// TIA Portal project "HEAT-1-CADIZ-V16" (V20)

(* hardware
DEVICE "S7-1200 station_1"  S7-1200 Station
   slot 0: "Rack_0"  S7-1200 Rack  Rack  V1.0
   slot 1: "PLC_1"  CPU 1214FC DC/DC/RLY  6ES7 214-1HF40-0XB0  V4.6
   slot 2: "DI 16x24VDC_1"  6ES7 221-1BH32-0XB0  V2.0
   slot 3: "DQ 16xRelay_1"  SM 1222 DQ16 x relay  6ES7 222-1HH32-0XB0  V2.0
   slot 4: "F-DI 8/16x24VDC_1"  SM 1226 F-DI8/16 x 24VDC  6ES7 226-6BA32-0XB0  V2.0
   slot 5: "F-DI 8/16x24VDC_2"  SM 1226 F-DI8/16 x 24VDC  6ES7 226-6BA32-0XB0  V2.0
   slot 6: "F-DQ 4x24VDC_1"  SM 1226 F-DQ4 x 24VDC  6ES7 226-6DA32-0XB0  V2.0
DEVICE "GSD device_1"  GSD.Device.PN
   slot 0: "Rack"  Rack  V1.0
   slot 0: "KRC5"  KUKA.PROFINET 6.0  0x300  V6.0
      slot 0: "KUKA.PROFINET 6.0"  KUKA.PROFINET 6.0
      slot 1: "Interface1"  Interface1
         slot 1: "Port001(XF3)"  Port001(XF3)
         slot 2: "Port002(XF4)"  Port002(XF4)
         slot 3: "Port003(XF5)"  Port003(XF5)
         slot 4: "Port004(XF6)"  Port004(XF6)
   slot 1: "64 safe digital in- and outputs (2.4)_1"  64 safe digital in- and outputs (2.4)  KUKADevF64_2.4
      slot 0: "64 safe digital in- and outputs (2.4)"  64 safe digital in- and outputs (2.4)
   slot 2: "512 digital in- and outputs_1"  512 digital in- and outputs  KUKA Device IO512
      slot 0: "512 digital in- and outputs"  512 digital in- and outputs
DEVICE "HMI_1"  KTP1200 Basic PN
   slot 0: "HMI_1"  KTP1200 Basic PN  6AV2 123-2MB03-0AX0  17.0.0.0
   slot 1: "HMI_RT_1"  KTP1200 Basic PN  6AV2 123-2MB03-0AX0  17.0.0.0
   slot 5: "HMI_1.IE_CP_1"  PROFINET Interface  17.0.0.0
      slot 1: "PROFINET Interface_1"  PROFINET Interface
         slot 1: "Port_1"  Port
DEVICE "ET 200SP station_2"  ET 200SP-Station
   slot 0: "Rack_0"  Rack  6ES5 710-8MAx1
   slot 0: "islaparking"  IM 155-6 PN ST  6ES7 155-6AU01-0BN0  V4.2
   slot 1: "DI 16x24VDC ST_1"  DI 16x24VDC ST  6ES7 131-6BH01-0BA0  V0.0
      slot 1: "DI 16x24VDC ST_1"  DI 16x24VDC ST
   slot 2: "DI 8x24VDC ST_1"  DI 8x24VDC ST  6ES7 131-6BF01-0BA0  V0.0
      slot 1: "DI 8x24VDC ST_1"  DI 8x24VDC ST
   slot 3: "DQ 16x24VDC/0.5A ST_1"  DQ 16x24VDC/0.5A ST  6ES7 132-6BH01-0BA0  V0.0
      slot 1: "DQ 16x24VDC/0.5A ST_1"  DQ 16x24VDC/0.5A ST
   slot 4: "DQ 8x24VDC/0.5A ST_1"  DQ 8x24VDC/0.5A ST  6ES7 132-6BF01-0BA0  V0.0
      slot 1: "DQ 8x24VDC/0.5A ST_1"  DQ 8x24VDC/0.5A ST
   slot 5: "Server module_1"  Server module  6ES7 193-6PA00-0AA0  V1.1
      slot 1: "Server module_1"  Server module
   slot 127: "BA 2xRJ45"  BA 2xRJ45  6ES7 193-6AR00-0AA0  V0.0
      slot 1: "Port_1"  X1 P1R  6ES7 193-6AR00-0AA0  V0.0
      slot 2: "Port_2"  X1 P2R  6ES7 193-6AR00-0AA0  V0.0
DEVICE "ET 200SP station_1"  ET 200SP-Station
   slot 0: "Rack_0"  Rack  6ES5 710-8MAx1
   slot 0: "islarobot"  IM 155-6 PN ST  6ES7 155-6AU01-0BN0  V4.2
   slot 1: "DI 16x24VDC ST_1"  DI 16x24VDC ST  6ES7 131-6BH01-0BA0  V0.0
      slot 1: "DI 16x24VDC ST_1"  DI 16x24VDC ST
   slot 2: "DI 8x24VDC ST_1"  DI 8x24VDC ST  6ES7 131-6BF01-0BA0  V0.0
      slot 1: "DI 8x24VDC ST_1"  DI 8x24VDC ST
   slot 3: "DQ 16x24VDC/0.5A ST_1"  DQ 16x24VDC/0.5A ST  6ES7 132-6BH01-0BA0  V0.0
      slot 1: "DQ 16x24VDC/0.5A ST_1"  DQ 16x24VDC/0.5A ST
   slot 4: "DQ 8x24VDC/0.5A ST_1"  DQ 8x24VDC/0.5A ST  6ES7 132-6BF01-0BA0  V0.0
      slot 1: "DQ 8x24VDC/0.5A ST_1"  DQ 8x24VDC/0.5A ST
   slot 5: "Server module_1"  Server module  6ES7 193-6PA00-0AA0  V1.1
      slot 1: "Server module_1"  Server module
   slot 127: "BA 2xRJ45"  BA 2xRJ45  6ES7 193-6AR00-0AA0  V0.0
      slot 1: "Port_1"  X1 P1R  6ES7 193-6AR00-0AA0  V0.0
      slot 2: "Port_2"  X1 P2R  6ES7 193-6AR00-0AA0  V0.0
DEVICE "GSD device_2"  GSD.Device.PN
   slot 0: "Rack"  Rack  V1.0
   slot 0: "CPX"  CPX Rev 50  TN 197330
      slot 0: "CPX Rev 50"  CPX Rev 50
      slot 1: "PN-IO Interface"  PN-IO Interface
         slot 1: "Port 1"  Port 1
         slot 2: "Port 2"  Port 2
   slot 1: "FB43 PNIO Module_1"  FB43 PNIO Module  TN 8110369, CPX-FB43
      slot 0: "FB43 PNIO Module"  FB43 PNIO Module
   slot 2: "MPAL DIL 4 [32DO]_1"  MPAL DIL 4 [32DO]
      slot 0: "MPAL DIL 4 [32DO]"  MPAL DIL 4 [32DO]
DEVICE "ET 200SP station_3"  ET 200SP-Station
   slot 0: "Rack_0"  Rack  6ES5 710-8MAx1
   slot 0: "sistemadeagua"  IM 155-6 PN ST  6ES7 155-6AU01-0BN0  V4.2
   slot 1: "DI 8x24VDC ST_1"  DI 8x24VDC ST  6ES7 131-6BF01-0BA0  V0.0
      slot 1: "DI 8x24VDC ST_1"  DI 8x24VDC ST
   slot 2: "DQ 8x24VDC/0.5A ST_1"  DQ 8x24VDC/0.5A ST  6ES7 132-6BF01-0BA0  V0.0
      slot 1: "DQ 8x24VDC/0.5A ST_1"  DQ 8x24VDC/0.5A ST
   slot 3: "AI 4xU/I 2-wire ST_1"  AI 4xU/I 2-wire ST  6ES7 134-6HD01-0BA1  V2.0
      slot 1: "AI 4xU/I 2-wire ST_1"  AI 4xU/I 2-wire ST
   slot 4: "Server module_1"  Server module  6ES7 193-6PA00-0AA0  V1.1
      slot 1: "Server module_1"  Server module
   slot 127: "BA 2xRJ45"  BA 2xRJ45  6ES7 193-6AR00-0AA0  V0.0
      slot 1: "Port_1"  X1 P1R  6ES7 193-6AR00-0AA0  V0.0
      slot 2: "Port_2"  X1 P2R  6ES7 193-6AR00-0AA0  V0.0
*)

// ===== PLC "PLC_1"  CPU 1214FC DC/DC/RLY =====

VAR_GLOBAL   // PLC tag table "Default tag table"
   "RES1 (reservado)" AT %Q500.0 : Bool;
   "eStopButtonCabinet" AT %I40.0 : Bool;   // Emergency-Stop cabinet — 1oo2 result
   "eStopButtonTank" AT %I40.1 : Bool;   // Emergency-Stop tank — 1oo2 result
   "eStopButtonTankPartnerCh" AT %I41.1 : Bool;   // partner channel 1oo2 — do not use
   "eStopButtonWaterSystem" AT %I40.2 : Bool;   // Emergency-Stop water system — 1oo2 result
   "eStopButtonWaterSystemPartnerCh" AT %I41.2 : Bool;   // partner channel 1oo2 — do not use
   "eStopButtonHmiPanel" AT %I40.3 : Bool;   // Emergency-Stop HMI panel — 1oo2 result
   "eStopButtonHmiPanelPartnerCh" AT %I41.3 : Bool;   // partner channel 1oo2 — do not use
   "eStopButtonLightCurtain1" AT %I40.4 : Bool;   // Emergency-Stop light curtain 1 — 1oo2 resul
   "eStopButtonLightCurtain1PartnerCh" AT %I41.4 : Bool;   // partner channel 1oo2 — do not use
   "eStopButtonDoor" AT %I40.5 : Bool;   // Emergency-Stop Door — 1oo2 result
   "eStopButtonDoorPartnerCh" AT %I41.5 : Bool;   // partner channel 1oo2 — do not use
   "lightCurtain1Ossd1" AT %I50.0 : Bool;   // Z2 – LC 1 OSSD 1 (receiver)
   "lightCurtain1Ossd2" AT %I51.0 : Bool;   // Z2 – LC 1 OSSD 2 (receiver)
   "lightCurtain3Ossd1" AT %I50.1 : Bool;   // Z2 – LC 3 OSSD 1 (receiver)
   "lightCurtain3Ossd2" AT %I51.1 : Bool;   // Z2 – LC 3 OSSD 2 (receiver)
   "lightCurtain6Ossd1" AT %I50.2 : Bool;   // Z2 – LC 6 OSSD 1 (receiver)
   "lightCurtain6Ossd2" AT %I51.2 : Bool;   // Z2 – LC 6 OSSD 2 (receiver)
   "enableAccessReqSelector" AT %I50.3 : Bool;   // Rotary selector – enabless request access
   "DoorClosedCh1" AT %I50.6 : Bool;   // Safety door closed interlock – contact 1
   "resetDoorButton" AT %I50.7 : Bool;   // Reset push‑button
   "SAF_DOOR_CLSD_CH2" AT %I51.6 : Bool;   // Safety door closed interlock – contact 2
   "SAF_DOOR_UNLOCK_CH1" AT %Q60.0 : Bool;   // Unlock safety door – redundant output 1
   "SAF_GATE_UNLOCK_CH2" AT %Q60.2 : Bool;   // Unlock safety door – redundant output 2
   "IND_RESET_LAMP" AT %Q10.0 : Bool;   // Reset indicator lamp
   "IND_STATUS_LAMP" AT %Q10.1 : Bool;   // System-status pilot light
   "CMD_PRESS_EXH_VALVE" AT %Q11.0 : Bool;   // Pressure/exhaust solenoid-valve command
   "STS_RECIRC_PUMP" AT %I20.0 : Bool;   // Recirculation-pump feedback
   "STS_TRANSFER_PUMP" AT %I20.1 : Bool;   // Transfer-pump feedback
   "ALM_UV_FILTER" AT %I20.2 : Bool;   // UV-filter fault alarm
   "ALM_PIT_LVL_LOW" AT %I20.3 : Bool;   // Sump low-level alarm
   "ALM_TANK_LVL_LOW" AT %I20.4 : Bool;   // Tank low-level alarm
   "STS_TANK_FILLING" AT %I20.5 : Bool;   // Tank filling status
   "STS_TANK_DRAINING" AT %I20.6 : Bool;   // Tank draining status
   "MODE_WATER_AUTO" AT %Q30.3 : Bool;   // CONMUTADOR AUTO
   "IND_BEACON2_GREEN" AT %Q30.4 : Bool;   // Beacon 2 – green
   "IND_BEACON2_RED" AT %Q30.5 : Bool;   // Beacon 2 – red
   "robotPresenceSignalZone1" AT %I500.0 : Bool;
   "robotPresenceSignalZone2" AT %I500.1 : Bool;
   "robotPresenceSignalZone3" AT %I500.2 : Bool;
   "eStopButtonCabinetPartnerCh" AT %I41.0 : Bool;   // partner channel 1oo2 — do not use
   "lightCurtain2Ossd1" AT %I300.0 : Bool;
   "lightCurtain2Ossd2" AT %I301.0 : Bool;
   "eStopButtonIslandRightPartner" AT %I301.1 : Bool;
   "lightCurtain4Ossd1" AT %I350.0 : Bool;
   "eStopButtonIslandLeft" AT %I350.1 : Bool;
   "lightCurtain5Ossd1" AT %I350.2 : Bool;
   "eStopButtonIslandLefttPartner" AT %I350.3 : Bool;   // partner channel 1oo2 — do not use
   "lightCurtain4Ossd2" AT %I350.4 : Bool;
   "lightCurtain5Ossd2" AT %I350.6 : Bool;
   "accessReqButtonZone2" AT %I51.4 : Bool;   // Illuminated push-button – access request for zone 2
   "accessReqButtonZone3" AT %I51.5 : Bool;   // Illuminated push-button – access request for zone 3
   "accessReqButtonZone1" AT %I51.3 : Bool;   // Illuminated push-button – access request for zone 1
   "eStopButtonIslandRight" AT %I300.1 : Bool;
   "NHE – E‑Stop externo  NO pulsado" AT %Q500.1 : Bool;
   "BS – Puerta cerrada" AT %Q500.2 : Bool;
   "QBS – Ack puerta" AT %Q500.3 : Bool;
   "SHS1 – Stop 1" AT %Q500.4 : Bool;
   "SHS2 – Stop 2" AT %Q500.5 : Bool;
   "RES6" AT %Q500.6 : Bool;
   "RES7" AT %Q500.7 : Bool;
   "US2 – 24 V US2" AT %Q501.0 : Bool;
   "SBH – Safe Op Stop" AT %Q501.1 : Bool;
   "RES11" AT %Q501.2 : Bool;
   "RES12" AT %Q501.3 : Bool;
   "RES13" AT %Q501.4 : Bool;
   "RES14" AT %Q501.5 : Bool;
   "RES15" AT %Q501.6 : Bool;
   "SPA – Power‑down Ack" AT %Q501.7 : Bool;
   "resetHmiButton" AT %I51.7 : Bool;
   "Tag_1" AT %M200.0 : Bool;
   "Tag_2" AT %M201.0 : Bool;
   "Tag_3" AT %M500.1 : Bool;
   "Tag_4" AT %M755.5 : Bool;
   "V5" AT %Q0.4 : Bool;   // Biestable_B_RETROCESO
   "ABRIR_TAPA_PEPA" AT %Q170.2 : Bool;
   "CERRAR_TAPA_PEPA" AT %Q170.3 : Bool;
   "ABRIR_TAPA_INMERSION" AT %Q170.4 : Bool;
   "CERRAR_TAPA_INMERSION" AT %Q170.5 : Bool;
   "ABRIR_TAPA_MARCADOR" AT %Q170.6 : Bool;
   "CERRAR_TAPA_MARCADOR" AT %Q170.7 : Bool;
   "ABRIR_TAPA_PERFILOMETRO" AT %Q171.0 : Bool;
   "CERRAR_TAPA_PERFILOMETRO" AT %Q171.1 : Bool;
   "V6" AT %Q0.5 : Bool;   // Biestable_A_AVANCE
   "V7" AT %Q0.6 : Bool;
   "V8" AT %Q0.7 : Bool;
   "moveCode_00" AT %Q616.0 : Bool;
   "goTrigger" AT %Q622.0 : Bool;
   "baseReqId_00" AT %Q620.0 : Bool;
   "baseReqId_01" AT %Q620.1 : Bool;
   "baseReqId_02" AT %Q620.2 : Bool;
   "baseReqId_03" AT %Q620.3 : Bool;
   "baseReqId_04" AT %Q620.4 : Bool;
   "baseReqId_05" AT %Q620.5 : Bool;
   "baseReqId_06" AT %Q620.6 : Bool;
   "baseReqId_07" AT %Q620.7 : Bool;
   "baseReqId_08" AT %Q621.0 : Bool;
   "baseReqId_09" AT %Q621.1 : Bool;
   "baseReqId_10" AT %Q621.2 : Bool;
   "baseReqId_11" AT %Q621.3 : Bool;
   "baseReqId_12" AT %Q621.4 : Bool;
   "baseReqId_13" AT %Q621.5 : Bool;
   "baseReqId_14" AT %Q621.6 : Bool;
   "baseReqId_15" AT %Q621.7 : Bool;
   "moveCode_01" AT %Q616.1 : Bool;
   "moveCode_02" AT %Q616.2 : Bool;
   "moveCode_03" AT %Q616.3 : Bool;
   "moveCode_04" AT %Q616.4 : Bool;
   "moveCode_05" AT %Q616.5 : Bool;
   "moveCode_06" AT %Q616.6 : Bool;
   "moveCode_07" AT %Q616.7 : Bool;
   "moveCode_08" AT %Q617.0 : Bool;
   "moveCode_09" AT %Q617.1 : Bool;
   "moveCode_10" AT %Q617.2 : Bool;
   "moveCode_11" AT %Q617.3 : Bool;
   "moveCode_12" AT %Q617.4 : Bool;
   "moveCode_13" AT %Q617.5 : Bool;
   "moveCode_14" AT %Q617.6 : Bool;
   "moveCode_15" AT %Q617.7 : Bool;
   "toolNo_00" AT %I625.0 : Bool;
   "toolNo_01" AT %I625.1 : Bool;
   "toolNo_02" AT %I625.2 : Bool;
   "toolNo_03" AT %I625.3 : Bool;
   "toolNo_04" AT %I625.4 : Bool;
   "toolNo_05" AT %I625.5 : Bool;
   "toolNo_06" AT %I625.6 : Bool;
   "toolNo_07" AT %I625.7 : Bool;
   "baseNo_00" AT %I626.0 : Bool;
   "baseNo_01" AT %I626.1 : Bool;
   "baseNo_02" AT %I626.2 : Bool;
   "baseNo_03" AT %I626.3 : Bool;
   "baseNo_04" AT %I626.4 : Bool;
   "baseNo_05" AT %I626.5 : Bool;
   "baseNo_06" AT %I626.6 : Bool;
   "baseNo_07" AT %I626.7 : Bool;
   "toolNoByte" AT %IB625 : Byte;
   "baseNoByte" AT %IB626 : Byte;
   "programReqId_00" AT %Q623.0 : Bool;
   "programReqId_01" AT %Q623.1 : Bool;
   "programReqId_02" AT %Q623.2 : Bool;
   "programReqId_03" AT %Q623.3 : Bool;
   "programReqId_04" AT %Q623.4 : Bool;
   "programReqId_05" AT %Q623.5 : Bool;
   "programReqId_06" AT %Q623.6 : Bool;
   "programReqId_07" AT %Q623.7 : Bool;
   "programReqId_08" AT %Q624.0 : Bool;
   "programReqId_09" AT %Q624.1 : Bool;
   "programReqId_10" AT %Q624.2 : Bool;
   "programReqId_11" AT %Q624.3 : Bool;
   "programReqId_12" AT %Q624.4 : Bool;
   "programReqId_13" AT %Q624.5 : Bool;
   "programReqId_14" AT %Q624.6 : Bool;
   "programReqId_15" AT %Q624.7 : Bool;
   "programReqId" AT %QW623 : Word;
   "PRUEBA_4" AT %Q4.4 : Bool;
   "PRUEBA_5" AT %Q4.5 : Bool;
   "PRUEBA_JOAQUIN" AT %Q4.0 : Bool;
   "PRUEBA_6" AT %Q4.6 : Bool;
   "PRUEBA_7" AT %Q4.7 : Bool;
   "cancelGo" AT %Q625.0 : Bool;
   "pauseGo" AT %Q625.1 : Bool;
   "resumeGo" AT %Q625.2 : Bool;
   "kukaCmdSafeForChange" AT %I624.4 : Bool;
   "cancelAck" AT %I624.5 : Bool;
   "pauseAck" AT %I624.6 : Bool;
   "resumeAck" AT %I624.7 : Bool;
END_VAR

VAR_GLOBAL   // PLC tag table "Robot Jog"
   "tcpTargetX_01" AT %Q600.1 : Bool;
   "tcpTargetX_02" AT %Q600.2 : Bool;
   "tcpTargetX_03" AT %Q600.3 : Bool;
   "tcpTargetX_04" AT %Q600.4 : Bool;
   "tcpTargetX_05" AT %Q600.5 : Bool;
   "tcpTargetX_08" AT %Q601.0 : Bool;
   "tcpTargetX_16" AT %Q602.0 : Bool;
   "tcpTargetX_17" AT %Q602.1 : Bool;
   "tcpTargetX_06" AT %Q600.6 : Bool;
   "tcpTargetX_07" AT %Q600.7 : Bool;
   "tcpTargetX_09" AT %Q601.1 : Bool;
   "tcpTargetX_10" AT %Q601.2 : Bool;
   "tcpTargetX_11" AT %Q601.3 : Bool;
   "tcpTargetX_12" AT %Q601.4 : Bool;
   "tcpTargetX_13" AT %Q601.5 : Bool;
   "tcpTargetX_14" AT %Q601.6 : Bool;
   "tcpTargetX_15" AT %Q601.7 : Bool;
   "tcpTargetX_18" AT %Q602.2 : Bool;
   "tcpTargetX_19" AT %Q602.3 : Bool;
   "tcpTargetX_20" AT %Q602.4 : Bool;
   "tcpTargetX_21" AT %Q602.5 : Bool;
   "tcpTargetX_22" AT %Q602.6 : Bool;
   "tcpTargetX_23" AT %Q602.7 : Bool;
   "tcpTargetX_24" AT %Q603.0 : Bool;
   "tcpTargetX_25" AT %Q603.1 : Bool;
   "tcpTargetX_26" AT %Q603.2 : Bool;
   "tcpTargetX_27" AT %Q603.3 : Bool;
   "tcpTargetX_28" AT %Q603.4 : Bool;
   "tcpTargetX_29" AT %Q603.5 : Bool;
   "tcpTargetX_30" AT %Q603.6 : Bool;
   "tcpTargetX_31" AT %Q603.7 : Bool;
   "tcpTargetY_00" AT %Q604.0 : Bool;
   "tcpTargetY_01" AT %Q604.1 : Bool;
   "tcpTargetY_02" AT %Q604.2 : Bool;
   "tcpTargetY_03" AT %Q604.3 : Bool;
   "tcpTargetY_04" AT %Q604.4 : Bool;
   "tcpTargetY_05" AT %Q604.5 : Bool;
   "tcpTargetY_06" AT %Q604.6 : Bool;
   "tcpTargetY_07" AT %Q604.7 : Bool;
   "tcpTargetY_08" AT %Q605.0 : Bool;
   "tcpTargetY_09" AT %Q605.1 : Bool;
   "tcpTargetY_10" AT %Q605.2 : Bool;
   "tcpTargetY_11" AT %Q605.3 : Bool;
   "tcpTargetY_12" AT %Q605.4 : Bool;
   "tcpTargetY_13" AT %Q605.5 : Bool;
   "tcpTargetY_14" AT %Q605.6 : Bool;
   "tcpTargetY_15" AT %Q605.7 : Bool;
   "tcpTargetY_16" AT %Q606.0 : Bool;   // $IN[49]
   "tcpTargetY_17" AT %Q606.1 : Bool;   // $IN[50]
   "tcpTargetY_18" AT %Q606.2 : Bool;   // $IN[51]
   "tcpTargetY_19" AT %Q606.3 : Bool;   // true
   "tcpTargetY_20" AT %Q606.4 : Bool;
   "tcpTargetY_21" AT %Q606.5 : Bool;   // true
   "tcpTargetY_22" AT %Q606.6 : Bool;   // true
   "tcpTargetY_23" AT %Q606.7 : Bool;   // true
   "tcpTargetY_24" AT %Q607.0 : Bool;   // true
   "tcpTargetY_25" AT %Q607.1 : Bool;   // true
   "tcpTargetY_26" AT %Q607.2 : Bool;   // true
   "tcpTargetY_27" AT %Q607.3 : Bool;
   "tcpTargetY_28" AT %Q607.4 : Bool;
   "tcpTargetY_29" AT %Q607.5 : Bool;
   "tcpTargetY_30" AT %Q607.6 : Bool;
   "tcpTargetY_31" AT %Q607.7 : Bool;
   "tcpTargetZ_00" AT %Q608.0 : Bool;
   "tcpTargetZ_01" AT %Q608.1 : Bool;
   "tcpTargetZ_02" AT %Q608.2 : Bool;
   "tcpTargetZ_03" AT %Q608.3 : Bool;
   "tcpTargetZ_04" AT %Q608.4 : Bool;
   "tcpTargetZ_05" AT %Q608.5 : Bool;
   "tcpTargetZ_06" AT %Q608.6 : Bool;
   "tcpTargetZ_07" AT %Q608.7 : Bool;
   "tcpTargetZ_08" AT %Q609.0 : Bool;
   "tcpTargetZ_09" AT %Q609.1 : Bool;
   "tcpTargetZ_10" AT %Q609.2 : Bool;
   "tcpTargetZ_11" AT %Q609.3 : Bool;
   "tcpTargetZ_12" AT %Q609.4 : Bool;
   "tcpTargetZ_13" AT %Q609.5 : Bool;
   "tcpTargetZ_14" AT %Q609.6 : Bool;
   "tcpTargetZ_15" AT %Q609.7 : Bool;
   "tcpTargetZ_16" AT %Q610.0 : Bool;
   "tcpTargetZ_17" AT %Q610.1 : Bool;
   "tcpTargetZ_18" AT %Q610.2 : Bool;
   "tcpTargetZ_19" AT %Q610.3 : Bool;
   "tcpTargetZ_20" AT %Q610.4 : Bool;
   "tcpTargetZ_21" AT %Q610.5 : Bool;
   "tcpTargetZ_22" AT %Q610.6 : Bool;
   "tcpTargetZ_23" AT %Q610.7 : Bool;
   "tcpTargetZ_24" AT %Q611.0 : Bool;
   "tcpTargetZ_25" AT %Q611.1 : Bool;
   "tcpTargetZ_26" AT %Q611.2 : Bool;
   "tcpTargetZ_27" AT %Q611.3 : Bool;
   "tcpTargetZ_28" AT %Q611.4 : Bool;
   "tcpTargetZ_29" AT %Q611.5 : Bool;
   "tcpTargetZ_30" AT %Q611.6 : Bool;
   "tcpTargetZ_31" AT %Q611.7 : Bool;
   "e1Target_00" AT %Q612.0 : Bool;
   "e1Target_01" AT %Q612.1 : Bool;
   "e1Target_02" AT %Q612.2 : Bool;
   "e1Target_03" AT %Q612.3 : Bool;
   "e1Target_04" AT %Q612.4 : Bool;
   "e1Target_05" AT %Q612.5 : Bool;
   "e1Target_06" AT %Q612.6 : Bool;
   "e1Target_07" AT %Q612.7 : Bool;
   "e1Target_08" AT %Q613.0 : Bool;
   "e1Target_09" AT %Q613.1 : Bool;
   "e1Target_10" AT %Q613.2 : Bool;
   "e1Target_11" AT %Q613.3 : Bool;
   "e1Target_12" AT %Q613.4 : Bool;
   "e1Target_13" AT %Q613.5 : Bool;
   "e1Target_14" AT %Q613.6 : Bool;
   "e1Target_15" AT %Q613.7 : Bool;
   "e1Target_16" AT %Q614.0 : Bool;
   "e1Target_17" AT %Q614.1 : Bool;
   "e1Target_18" AT %Q614.2 : Bool;
   "e1Target_19" AT %Q614.3 : Bool;
   "e1Target_20" AT %Q614.4 : Bool;
   "e1Target_21" AT %Q614.5 : Bool;
   "e1Target_22" AT %Q614.6 : Bool;
   "e1Target_23" AT %Q614.7 : Bool;
   "e1Target_24" AT %Q615.0 : Bool;
   "e1Target_25" AT %Q615.1 : Bool;
   "e1Target_26" AT %Q615.2 : Bool;
   "e1Target_27" AT %Q615.3 : Bool;
   "e1Target_28" AT %Q615.4 : Bool;
   "e1Target_29" AT %Q615.5 : Bool;
   "e1Target_30" AT %Q615.6 : Bool;
   "e1Target_31" AT %Q615.7 : Bool;
   "e1Target_Word" AT %QD612 : DWord;
   "moveCodeKuka" AT %QW616 : Word;   // SIGNAL goTrrigger $IN[ 129]
   "rbDone" AT %I624.0 : Bool;   // SIGNAL rbDoneEdge $OUT[193]
   "x1Target_Word" AT %QD600 : DWord;
   "y1Target_Word" AT %QD604 : DWord;
   "z1Target_Word" AT %QD608 : DWord;
END_VAR

VAR_GLOBAL   // PLC tag table "Robot Position"
   "tcpPosIniX_00" AT %I632.0 : Bool;
   "tcpPosIniX_01" AT %I632.1 : Bool;
   "tcpPosIniX_02" AT %I632.2 : Bool;
   "tcpPosIniX_03" AT %I632.3 : Bool;
   "tcpPosIniX_04" AT %I632.4 : Bool;
   "tcpPosIniX_05" AT %I632.5 : Bool;
   "tcpPosIniX_06" AT %I632.6 : Bool;
   "tcpPosIniX_07" AT %I632.7 : Bool;
   "tcpPosIniX_08" AT %I633.0 : Bool;
   "tcpPosIniX_09" AT %I633.1 : Bool;
   "tcpPosIniX_10" AT %I633.2 : Bool;
   "tcpPosIniX_11" AT %I633.3 : Bool;
   "tcpPosIniX_12" AT %I633.4 : Bool;
   "tcpPosIniX_13" AT %I633.5 : Bool;
   "tcpPosIniX_14" AT %I633.6 : Bool;
   "tcpPosIniX_15" AT %I633.7 : Bool;
   "tcpPosIniX_16" AT %I634.0 : Bool;
   "tcpPosIniX_17" AT %I634.1 : Bool;
   "tcpPosIniX_18" AT %I634.2 : Bool;
   "tcpPosIniX_19" AT %I634.3 : Bool;
   "tcpPosIniX_20" AT %I634.4 : Bool;
   "tcpPosIniX_21" AT %I634.5 : Bool;
   "tcpPosIniX_22" AT %I634.6 : Bool;
   "tcpPosIniX_23" AT %I634.7 : Bool;
   "tcpPosIniX_24" AT %I635.0 : Bool;
   "tcpPosIniX_25" AT %I635.1 : Bool;
   "tcpPosIniX_26" AT %I635.2 : Bool;
   "tcpPosIniX_27" AT %I635.3 : Bool;
   "tcpPosIniX_28" AT %I635.4 : Bool;
   "tcpPosIniX_29" AT %I635.5 : Bool;
   "tcpPosIniX_30" AT %I635.6 : Bool;
   "tcpPosIniX_31" AT %I635.7 : Bool;
   "tcpPosIniY_00" AT %I636.0 : Bool;
   "tcpPosIniY_01" AT %I636.1 : Bool;
   "tcpPosIniY_02" AT %I636.2 : Bool;
   "tcpPosIniY_03" AT %I636.3 : Bool;
   "tcpPosIniY_04" AT %I636.4 : Bool;
   "tcpPosIniY_05" AT %I636.5 : Bool;
   "tcpPosIniY_06" AT %I636.6 : Bool;
   "tcpPosIniY_07" AT %I636.7 : Bool;
   "tcpPosIniY_08" AT %I637.0 : Bool;
   "tcpPosIniY_09" AT %I637.1 : Bool;
   "tcpPosIniY_10" AT %I637.2 : Bool;
   "tcpPosIniY_11" AT %I637.3 : Bool;
   "tcpPosIniY_12" AT %I637.4 : Bool;
   "tcpPosIniY_13" AT %I637.5 : Bool;
   "tcpPosIniY_14" AT %I637.6 : Bool;
   "tcpPosIniY_15" AT %I637.7 : Bool;
   "tcpPosIniY_16" AT %I638.0 : Bool;
   "tcpPosIniY_17" AT %I638.1 : Bool;
   "tcpPosIniY_18" AT %I638.2 : Bool;
   "tcpPosIniY_19" AT %I638.3 : Bool;
   "tcpPosIniY_20" AT %I638.4 : Bool;
   "tcpPosIniY_21" AT %I638.5 : Bool;
   "tcpPosIniY_22" AT %I638.6 : Bool;
   "tcpPosIniY_23" AT %I638.7 : Bool;
   "tcpPosIniY_24" AT %I639.0 : Bool;
   "tcpPosIniY_25" AT %I639.1 : Bool;
   "tcpPosIniY_26" AT %I639.2 : Bool;
   "tcpPosIniY_27" AT %I639.3 : Bool;
   "tcpPosIniY_28" AT %I639.4 : Bool;
   "tcpPosIniY_29" AT %I639.5 : Bool;
   "tcpPosIniY_30" AT %I639.6 : Bool;
   "tcpPosIniY_31" AT %I639.7 : Bool;
   "tcpPosIniZ_00" AT %I640.0 : Bool;
   "tcpPosIniZ_01" AT %I640.1 : Bool;
   "tcpPosIniZ_02" AT %I640.2 : Bool;
   "tcpPosIniZ_03" AT %I640.3 : Bool;
   "tcpPosIniZ_04" AT %I640.4 : Bool;
   "tcpPosIniZ_05" AT %I640.5 : Bool;
   "tcpPosIniZ_06" AT %I640.6 : Bool;
   "tcpPosIniZ_07" AT %I640.7 : Bool;
   "tcpPosIniZ_08" AT %I641.0 : Bool;
   "tcpPosIniZ_09" AT %I641.1 : Bool;
   "tcpPosIniZ_10" AT %I641.2 : Bool;
   "tcpPosIniZ_11" AT %I641.3 : Bool;
   "tcpPosIniZ_12" AT %I641.4 : Bool;
   "tcpPosIniZ_13" AT %I641.5 : Bool;
   "tcpPosIniZ_14" AT %I641.6 : Bool;
   "tcpPosIniZ_15" AT %I641.7 : Bool;
   "tcpPosIniZ_16" AT %I642.0 : Bool;
   "tcpPosIniZ_17" AT %I642.1 : Bool;
   "tcpPosIniZ_18" AT %I642.2 : Bool;
   "tcpPosIniZ_19" AT %I642.3 : Bool;
   "tcpPosIniZ_20" AT %I642.4 : Bool;
   "tcpPosIniZ_21" AT %I642.5 : Bool;
   "tcpPosIniZ_22" AT %I642.6 : Bool;
   "tcpPosIniZ_23" AT %I642.7 : Bool;
   "tcpPosIniZ_24" AT %I643.0 : Bool;
   "tcpPosIniZ_25" AT %I643.1 : Bool;
   "tcpPosIniZ_26" AT %I643.2 : Bool;
   "tcpPosIniZ_27" AT %I643.3 : Bool;
   "tcpPosIniZ_28" AT %I643.4 : Bool;
   "tcpPosIniZ_29" AT %I643.5 : Bool;
   "tcpPosIniZ_30" AT %I643.6 : Bool;
   "tcpPosIniZ_31" AT %I643.7 : Bool;
   "e1PosIni_00" AT %I644.0 : Bool;
   "e1PosIni_01" AT %I644.1 : Bool;
   "e1PosIni_02" AT %I644.2 : Bool;
   "e1PosIni_03" AT %I644.3 : Bool;
   "e1PosIni_04" AT %I644.4 : Bool;
   "e1PosIni_05" AT %I644.5 : Bool;
   "e1PosIni_06" AT %I644.6 : Bool;
   "e1PosIni_07" AT %I644.7 : Bool;
   "e1PosIni_08" AT %I645.0 : Bool;
   "e1PosIni_09" AT %I645.1 : Bool;
   "e1PosIni_10" AT %I645.2 : Bool;
   "e1PosIni_11" AT %I645.3 : Bool;
   "e1PosIni_12" AT %I645.4 : Bool;
   "e1PosIni_13" AT %I645.5 : Bool;
   "e1PosIni_14" AT %I645.6 : Bool;
   "e1PosIni_15" AT %I645.7 : Bool;
   "e1PosIni_16" AT %I646.0 : Bool;
   "e1PosIni_17" AT %I646.1 : Bool;
   "e1PosIni_18" AT %I646.2 : Bool;
   "e1PosIni_19" AT %I646.3 : Bool;
   "e1PosIni_20" AT %I646.4 : Bool;
   "e1PosIni_21" AT %I646.5 : Bool;
   "e1PosIni_22" AT %I646.6 : Bool;
   "e1PosIni_23" AT %I646.7 : Bool;
   "e1PosIni_24" AT %I647.0 : Bool;
   "e1PosIni_25" AT %I647.1 : Bool;
   "e1PosIni_26" AT %I647.2 : Bool;
   "e1PosIni_27" AT %I647.3 : Bool;
   "e1PosIni_28" AT %I647.4 : Bool;
   "e1PosIni_29" AT %I647.5 : Bool;
   "e1PosIni_30" AT %I647.6 : Bool;
   "e1PosIni_31" AT %I647.7 : Bool;
   "tcpPosFinX_00" AT %I648.0 : Bool;
   "tcpPosFinX_01" AT %I648.1 : Bool;
   "tcpPosFinX_02" AT %I648.2 : Bool;
   "tcpPosFinX_03" AT %I648.3 : Bool;
   "tcpPosFinX_04" AT %I648.4 : Bool;
   "tcpPosFinX_05" AT %I648.5 : Bool;
   "tcpPosFinX_06" AT %I648.6 : Bool;
   "tcpPosFinX_07" AT %I648.7 : Bool;
   "tcpPosFinX_08" AT %I649.0 : Bool;
   "tcpPosFinX_09" AT %I649.1 : Bool;
   "tcpPosFinX_10" AT %I649.2 : Bool;
   "tcpPosFinX_11" AT %I649.3 : Bool;
   "tcpPosFinX_12" AT %I649.4 : Bool;
   "tcpPosFinX_13" AT %I649.5 : Bool;
   "tcpPosFinX_14" AT %I649.6 : Bool;
   "tcpPosFinX_15" AT %I649.7 : Bool;
   "tcpPosFinX_16" AT %I650.0 : Bool;
   "tcpPosFinX_17" AT %I650.1 : Bool;
   "tcpPosFinX_18" AT %I650.2 : Bool;
   "tcpPosFinX_19" AT %I650.3 : Bool;
   "tcpPosFinX_20" AT %I650.4 : Bool;
   "tcpPosFinX_21" AT %I650.5 : Bool;
   "tcpPosFinX_22" AT %I650.6 : Bool;
   "tcpPosFinX_23" AT %I650.7 : Bool;
   "tcpPosFinX_24" AT %I651.0 : Bool;
   "tcpPosFinX_25" AT %I651.1 : Bool;
   "tcpPosFinX_26" AT %I651.2 : Bool;
   "tcpPosFinX_27" AT %I651.3 : Bool;
   "tcpPosFinX_28" AT %I651.4 : Bool;
   "tcpPosFinX_29" AT %I651.5 : Bool;
   "tcpPosFinX_30" AT %I651.6 : Bool;
   "tcpPosFinX_31" AT %I651.7 : Bool;
   "tcpPosFinY_00" AT %I652.0 : Bool;
   "tcpPosFinY_01" AT %I652.1 : Bool;
   "tcpPosFinY_02" AT %I652.2 : Bool;
   "tcpPosFinY_03" AT %I652.3 : Bool;
   "tcpPosFinY_04" AT %I652.4 : Bool;
   "tcpPosFinY_05" AT %I652.5 : Bool;
   "tcpPosFinY_06" AT %I652.6 : Bool;
   "tcpPosFinY_07" AT %I652.7 : Bool;
   "tcpPosFinY_08" AT %I653.0 : Bool;
   "tcpPosFinY_09" AT %I653.1 : Bool;
   "tcpPosFinY_10" AT %I653.2 : Bool;
   "tcpPosFinY_11" AT %I653.3 : Bool;
   "tcpPosFinY_12" AT %I653.4 : Bool;
   "tcpPosFinY_13" AT %I653.5 : Bool;
   "tcpPosFinY_14" AT %I653.6 : Bool;
   "tcpPosFinY_15" AT %I653.7 : Bool;
   "tcpPosFinY_16" AT %I654.0 : Bool;
   "tcpPosFinY_17" AT %I654.1 : Bool;
   "tcpPosFinY_18" AT %I654.2 : Bool;
   "tcpPosFinY_19" AT %I654.3 : Bool;
   "tcpPosFinY_20" AT %I654.4 : Bool;
   "tcpPosFinY_21" AT %I654.5 : Bool;
   "tcpPosFinY_22" AT %I654.6 : Bool;
   "tcpPosFinY_23" AT %I654.7 : Bool;
   "tcpPosFinY_24" AT %I655.0 : Bool;
   "tcpPosFinY_25" AT %I655.1 : Bool;
   "tcpPosFinY_26" AT %I655.2 : Bool;
   "tcpPosFinY_27" AT %I655.3 : Bool;
   "tcpPosFinY_28" AT %I655.4 : Bool;
   "tcpPosFinY_29" AT %I655.5 : Bool;
   "tcpPosFinY_30" AT %I655.6 : Bool;
   "tcpPosFinY_31" AT %I655.7 : Bool;
   "tcpPosE1_01" AT %I628.0 : Bool;
   "tcpPosE1_02" AT %I628.1 : Bool;
   "tcpPosE1_03" AT %I628.2 : Bool;
   "tcpPosE1_04" AT %I628.3 : Bool;
   "tcpPosE1_05" AT %I628.4 : Bool;
   "tcpPosE1_06" AT %I628.5 : Bool;
   "tcpPosE1_07" AT %I628.6 : Bool;
   "tcpPosE1_08" AT %I628.7 : Bool;
   "tcpPosE1_09" AT %I629.0 : Bool;
   "tcpPosE1_10" AT %I629.1 : Bool;
   "tcpPosE1_11" AT %I629.2 : Bool;
   "tcpPosE1_12" AT %I629.3 : Bool;
   "tcpPosE1_13" AT %I629.4 : Bool;
   "tcpPosE1_14" AT %I629.5 : Bool;
   "tcpPosE1_15" AT %I629.6 : Bool;
   "tcpPosE1_16" AT %I629.7 : Bool;
   "tcpPosE1_17" AT %I630.0 : Bool;
   "tcpPosE1_18" AT %I630.1 : Bool;
   "tcpPosE1_19" AT %I630.2 : Bool;
   "tcpPosE1_20" AT %I630.3 : Bool;
   "tcpPosE1_21" AT %I630.4 : Bool;
   "tcpPosE1_22" AT %I630.5 : Bool;
   "tcpPosE1_23" AT %I630.6 : Bool;
   "tcpPosE1_24" AT %I630.7 : Bool;
   "tcpPosE1_25" AT %I631.0 : Bool;
   "tcpPosE1_26" AT %I631.1 : Bool;
   "tcpPosE1_27" AT %I631.2 : Bool;
   "tcpPosE1_28" AT %I631.3 : Bool;
   "tcpPosE1_29" AT %I631.4 : Bool;
   "tcpPosE1_30" AT %I631.5 : Bool;
   "tcpPosE1_31" AT %I631.6 : Bool;
   "tcpPosE1_32" AT %I631.7 : Bool;
   "tcpPosIniX_rawLe32" AT %ID632 : DWord;
   "tcpPosIniY_rawLe32" AT %ID636 : DWord;
   "tcpPosIniZ_rawLe32" AT %ID640 : DWord;
   "tcpPosFinX_rawLe32" AT %ID648 : DWord;
   "tcpPosFinY_rawLe32" AT %ID652 : DWord;
   "e1_rawLe32" AT %ID628 : DWord;
   "e1PosIni_rawLe32" AT %ID644 : DWord;
   "tcpPosFinZ_rawLe32" AT %ID656 : DWord;
   "e1PosFin_rawLe32" AT %ID660 : DWord;
END_VAR

VAR_GLOBAL   // PLC tag table "Tool Change"
   "dockSensorToolInPosition" AT %I150.0 : Bool;   // DETECTOR_YUGO_LP
   "dockSensorCoverClosed" AT %I150.1 : Bool;   // TAPA_CERRADA_YUGO_LP
   "dockSensorCoverOpen" AT %I160.0 : Bool;   // TAPA_ABIERTA_YUGO_LP
   "dockValveV2UnlockOn" AT %Q171.2 : Bool;   // SOLTAR_HERRAMIENTA_YUGO_LP / CAMBIA A FALSE
   "dockValveCoverOpenOn" AT %Q170.0 : Bool;   // ABRIR_TAPA_YUGO_LP
   "dockValveCoverCloseOn" AT %Q170.1 : Bool;   // CERRAR_TAPA_YUGO_LP
   "robotSensorMpsUnlocked" AT %I200.0 : Bool;   // INTERCAMBIO_DESBLOQUEADO_LR
   "robotSensorMpsLocked" AT %I200.1 : Bool;   // INTERCAMBIO_BLOQUEADO_LR
   "robotSensorMpsCoupled" AT %I200.2 : Bool;   // HERRAMIENTA_PUESTA_LR /AL COLOCAR METAL
   "robotSensorMpsCtrlAirPressureOk" AT %I200.3 : Bool;   // PRESION_CORRECTA_LR
   "toolReqId_01" AT %Q618.1 : Bool;   // INKUKA_DETECTOR_HERRAMIENTA
   "toolReqId_02" AT %Q618.2 : Bool;   // INKUKA_TAPA_CERRADA_YUGO
   "toolReqId_03" AT %Q618.3 : Bool;   // INKUKA_TAPA_ABIERTA_YUGO
   "toolReqId_04" AT %Q618.4 : Bool;   // INKUKA_INTERCAMBIO_DESBLOQUEADO
   "toolReqId_05" AT %Q618.5 : Bool;   // INKUKA_INTERCAMBIO_BLOQUEADO
   "toolReqId_06" AT %Q618.6 : Bool;   // INKUKA_HERRAMIENTA_PUESTA /AL COLOCAR util met
   "toolReqId_07" AT %Q618.7 : Bool;
   "kukaCmdUnlockMps" AT %I624.1 : Bool;   // OUTKUKA_SOLTAR_HERRAMIENTA_YUGO
   "kukaCmdOpenCover" AT %I624.2 : Bool;   // OUTKUKA_ABRIR_TAPA_YUGO
   "kukaCmdCloseCover" AT %I624.3 : Bool;   // OUTKUKA_CERRAR_TAPA_YUGO
   "V1_B14_S2" AT %Q0.0 : Bool;   // Anticolision
   "V1_B12_S4" AT %Q0.1 : Bool;   // Mps Bloqueo SIL 2
   "V2_B14_S2" AT %Q0.2 : Bool;
   "V2_B12_S4" AT %Q0.3 : Bool;
   "toolReqId_00" AT %Q618.0 : Bool;
   "toolReqId_08" AT %Q619.0 : Bool;
   "toolReqId_09" AT %Q619.1 : Bool;
   "toolReqId_10" AT %Q619.2 : Bool;
   "toolReqId_11" AT %Q619.3 : Bool;
   "toolReqId_12" AT %Q619.4 : Bool;
   "toolReqId_13" AT %Q619.5 : Bool;
   "toolReqId_14" AT %Q619.6 : Bool;
   "toolReqId_15" AT %Q619.7 : Bool;
   "toolReqId" AT %QW618 : Word;
   "baseReqId" AT %QW620 : Word;
   "kukaFeedbackDockToolInPosition" AT %Q622.1 : Bool;
   "kukaFeedbackDockCoverClosed" AT %Q622.2 : Bool;
   "kukaFeedbackDockCoverOpen" AT %Q622.3 : Bool;
   "kukaFeedbackRobotMpsUnlocked" AT %Q622.4 : Bool;
   "kukaFeedbackRobotMpsLocked" AT %Q622.5 : Bool;
   "kukaFeedbackRobotMpsCoupled" AT %Q622.6 : Bool;
   "kukaFeedbackRobotMpsCtrlAirPressureOk" AT %Q622.7 : Bool;
END_VAR

VAR_GLOBAL   // PLC tag table "General"
   "ALM_PRESS_SENSOR" AT %I10.0 : Bool;   // Pressure-sensor alarm
   "CMD_TANK_FILL" AT %Q30.0 : Bool;   // LLENAR CUBA
   "CMD_TANK_DRAIN" AT %Q30.1 : Bool;   // VACIAR CUBA
   "RECIRCULACION" AT %Q30.2 : Bool;   // CONMUTADOR MANUAL / cambiado a recirculacion
END_VAR

TYPE "UDT_Dock"
   STRUCT
      Sensor : Struct
         CoverOpen : Bool;
         CoverClosed : Bool;
         ToolInPosition : Bool;
      END_STRUCT;
      Valve : Struct
         CoverOpenOn : Bool;
         CoverCloseOn : Bool;
         V2UnlockOn : Bool;
      END_STRUCT;
   END_STRUCT;
END_TYPE

TYPE "UDT_RobotMps"
   STRUCT
      Sensor : Struct
         Coupled : Bool;
         Locked : Bool;
         Unlocked : Bool;
         CtrlAirPressureOk : Bool;
      END_STRUCT;
   END_STRUCT;
END_TYPE

// folder: 10. System/DbsInstancia

DATA_BLOCK "InstKukaControlSeq"   // DB14
{ S7_Optimized_Access := 'TRUE' }
VERSION : 0.1
// stored: InstanceOfName KukaControlSeq
"KukaControlSeq"
BEGIN
END_DATA_BLOCK

DATA_BLOCK "InstSupervisorSeq"   // DB15
{ S7_Optimized_Access := 'TRUE' }
VERSION : 0.1
// stored: InstanceOfName SupervisorSeq
"SupervisorSeq"
BEGIN
END_DATA_BLOCK

DATA_BLOCK "InstSeqManager"   // DB16
{ S7_Optimized_Access := 'TRUE' }
VERSION : 0.1
// stored: InstanceOfName SeqManager
"SeqManager"
BEGIN
END_DATA_BLOCK

// folder: 10. System/DbsOpcUa

DATA_BLOCK "PlcStatus"   // DB4
{ S7_Optimized_Access := 'TRUE' }
VERSION : 0.1
   VAR
      "- FOR  KUKACONTROL-" : Bool;
      mode : Struct
         effective : UInt;
         ready : Bool;
      END_STRUCT;
      active : Struct
         baseId : UInt;
         toolId : UInt;
         profileId : UInt;
      END_STRUCT;
      exec : Struct
         ackSeq : UInt;
         accepted : Bool;
         busy : Bool;
         done : Bool;
         error : Bool;
         errorCode : UDInt;
         cancelAck : Bool;
         pauseAck : Bool;
         resumeAck : Bool;
         paused : Bool;
      END_STRUCT;
      pose : Struct
         tcpPosX_mm : LReal;
         tcpPosY_mm : LReal;
         tcpPosZ_mm : LReal;
         tcpOriA_deg : LReal;
         tcpOriB_deg : LReal;
         tcpOriC_deg : LReal;
         e1Pos_mm : LReal;
      END_STRUCT;
      teach : Struct
         startX_mm : LReal;
         startY_mm : LReal;
         startZ_mm : LReal;
         startE1_mm : LReal;
         startOk : Bool;
         endX_mm : LReal;
         endY_mm : LReal;
         endZ_mm : LReal;
         endE1_mm : LReal;
         endOk : Bool;
      END_STRUCT;
      "- FOR SUPERVISOR -" : Bool;
      heartbeatPlc : Bool;
      stepPlc : Int;
      plcOk : Bool;
      safetyOk : Bool;
      airOk : Bool;
      inspWaterOk : Bool;
      tankWaterOk : Bool;
      robotOk : Bool;
      acknowledge : Bool;
      carriageId : String;
      newCarriageId : Bool;
      idRunning : Bool;
      idOk : Bool;
      startUsReady : Bool;
      stopUsReady : Bool;
      paCheckReady : Bool;
      gainReady : Bool;
      tcgReady : Bool;
      idScan : String;
      pointOrigin : LReal;
      xSize : LReal;
      ySize : LReal;
      scanRefStart : Bool;
      scanInspStart : Bool;
      markRunning : Bool;
      markState : Bool;
      breakUs : Bool;
      unbreakUs : Bool;
      robotRescanning : Bool;
      acknowledgeError : Bool;
   END_VAR
BEGIN
END_DATA_BLOCK

DATA_BLOCK "KukaControlCmd"   // DB5
{ S7_Optimized_Access := 'TRUE' }
VERSION : 0.1
   VAR
      code : UInt;
      seq : UInt;
      tcpTargetX_mm : LReal;
      tcpTargetY_mm : LReal;
      tcpTargetZ_mm : LReal;
      e1Target : LReal;
      toolRequestId : UInt;
      baseRequestId : UInt;
      profileRequestId : UInt;
      vel_mms : LReal;
      index_mm : LReal;
      apo_mm : LReal;
      programRequestId : UInt;
      cancelGo : Bool;
      pauseGo : Bool;
      resumeGo : Bool;
      mode : Struct
         request : UInt;
         reqSeq : UInt;
      END_STRUCT;
   END_VAR
BEGIN
END_DATA_BLOCK

DATA_BLOCK "SupervisorCmd"   // DB6
{ S7_Optimized_Access := 'TRUE' }
VERSION : 0.1
   VAR
      heartbeatSupervisor : Bool;
      stepSupervisor : Int;
      supervisorOk : Bool;
      stateUs : Bool;
      reqCarriageId : Bool;
      reqId : Bool;
      pns : String;
      referencePart : String;
      endEffector : Int;
      utTech : UInt;
      teachReq : Bool;
      paCheckReq : Bool;
      tcgReq : Bool;
      startUsRunning : Bool;
      stopUsRunning : Bool;
      elemState : Bool;
      elemRunning : Bool;
      balState : Bool;
      balRunning : Bool;
      gainState : Bool;
      gainRunning : Bool;
      tcgInProgress : Bool;
      tcgNextStep : Bool;
      tcgState : Bool;
      reqRefPart : Bool;
      reqStopCycle : Bool;
      reqTcgAdj : Bool;
      scanRefState : Bool;
      scanRefRunning : Bool;
      reqPreEval : Bool;
      reqIdentificationState : Bool;
      scanInspState : Bool;
      scanInsprunning : Bool;
      reqMark : Bool;
      reqVerif : Bool;
      pointCoordinates : LReal;
      goBack : Bool;
      rescanning : Bool;
      errorMessage : String;
      errorOcurred : Bool;
      gainAdjustmentReq : Bool;
   END_VAR
BEGIN
END_DATA_BLOCK

// folder: 10. System/Utilities

DATA_BLOCK "ConstantsDB"   // DB37
{ S7_Optimized_Access := 'TRUE' }
VERSION : 0.1
BEGIN
END_DATA_BLOCK

// folder: 20. Robot Services/AutoExt

DATA_BLOCK "instAutoExtSeq"   // DB7
{ S7_Optimized_Access := 'TRUE' }
VERSION : 0.1
// stored: InstanceOfName AutoExtSeq
"AutoExtSeq"
BEGIN
END_DATA_BLOCK

// folder: 20. Robot Services/DbsInstancia

DATA_BLOCK "InstTcpJogging"   // DB2
{ S7_Optimized_Access := 'TRUE' }
VERSION : 0.1
// stored: InstanceOfName TcpJogging
"TcpJogging"
BEGIN
END_DATA_BLOCK

DATA_BLOCK "ToolChange_DB"   // DB8
{ S7_Optimized_Access := 'TRUE' }
VERSION : 0.1
// stored: InstanceOfName ToolChange
"ToolChange"
BEGIN
END_DATA_BLOCK

DATA_BLOCK "TcpPoseDecoderLe32_DB"   // DB10
{ S7_Optimized_Access := 'TRUE' }
VERSION : 0.1
// stored: InstanceOfName TcpPoseDecoderLe32
"TcpPoseDecoderLe32"
BEGIN
END_DATA_BLOCK

DATA_BLOCK "InstTcpTarget"   // DB13
{ S7_Optimized_Access := 'TRUE' }
VERSION : 0.1
// stored: InstanceOfName TcpTarget
"TcpTarget"
BEGIN
END_DATA_BLOCK

// folder: 30. Safety

DATA_BLOCK "InstMainSafety"   // DB1, F_DB
{ S7_Optimized_Access := 'TRUE' }
NAME : FUSI
VERSION : 0.1
// stored: InstanceOfName MainSafety
"MainSafety"
BEGIN
END_DATA_BLOCK

DATA_BLOCK "SafetyRobotDb"   // DB3, F_DB
{ S7_Optimized_Access := 'TRUE' }
VERSION : 0.1
BEGIN
END_DATA_BLOCK

// folder: Eliminar

DATA_BLOCK "DB_Supervisor"   // DB9
{ S7_Optimized_Access := 'TRUE' }
VERSION : 0.1
   VAR
      Common : Struct
         plc_ok : Bool;
         supervisor_ok : Bool;
         system_ok : Bool;
         safety_ok : Bool;
         air_ok : Bool;
         insp_water_ok : Bool;
         tank_water_ok : Bool;
         robot_ok : Bool;
         step_plc : Int;
         step_supervisor : Int;
         error : Bool;
         reset_req : Bool;
      END_STRUCT;
      Identification : Struct   // pag 2
         carriage_id_req : Bool;   // Sup->PLC
         new_carriage_id : Bool;   // PLC->Sup
         id_req : Bool;   // Sup->PLC
         id_running : Bool;   // PLC->Sup
         id_ok : Bool;   // PLC->Sup
         teach_req : Bool;   // Sup->PLC
         system_ok : Bool;   // PLC->Sup (parte de id_ok)
         pa_check_req : Bool;   // Sup->PLC
         tcg_req : Bool;   // Sup->PLC
      END_STRUCT;
      Teaching : Struct   // pag 3
         teach_ready : Bool;   // PLC->Sup
         teach_running : Bool;   // Sup->PLC
         teach_state : Bool;   // Sup->PLC
         jump_start_us : Bool;   // PLC->Sup
      END_STRUCT;
      StartUs : Struct   // pag 4
         start_us_ready : Bool;   // PLC->Sup
         start_us_running : Bool;   // Sup->PLC
         start_us_state : Bool;   // Sup->PLC
      END_STRUCT;
      PACheck : Struct   // pag 5
         pa_check_ready : Bool;   // PLC->Sup
         elem_running : Bool;   // Sup->PLC
         elem_state : Bool;   // Sup->PLC
         bal_running : Bool;   // Sup->PLC
         bal_state : Bool;   // Sup->PLC
      END_STRUCT;
      Gain : Struct
         gain_ready : Bool;
         gain_running : Bool;
         gain_state : Bool;
      END_STRUCT;
      TCG_Check : Struct
         tcg_ready : Bool;
         tcg_running : Bool;
         tcg_next_step : Bool;
         jump_acq_ref : Bool;
         jump_tcg_adj : Bool;
      END_STRUCT;
      TCG_Adjust : Struct
         tcg_ready : Bool;
         jump_ref_acq : Bool;
      END_STRUCT;
      RefScan_Acq : Struct
         scan_ref_ready : Bool;
         scan_ref_running : Bool;
      END_STRUCT;
      InspScan : Struct
         scan_insp_ready : Bool;
         scan_insp_running : Bool;
         scan_insp_state : Bool;
         jump_ref_insp : Bool;
      END_STRUCT;
      RefScan_Verif : Struct
         scan_ref_ready : Bool;
         scan_ref_running : Bool;
         jump_start : Bool;
      END_STRUCT;
      Marking : Struct
         mark_req : Bool;
         mark_running : Bool;
         mark_state : Bool;
         jump_start : Bool;
         point_coordinates : Struct
            x : Real;
            y : Real;
            z : Real;
            "a" : Real;
            "b" : Real;
            c : Real;
         END_STRUCT;
      END_STRUCT;
   END_VAR
BEGIN
END_DATA_BLOCK

// folder: 10. System

FUNCTION_BLOCK "SeqManager"   // FB20, LAD
{ S7_Optimized_Access := 'TRUE' }
VERSION : 0.1
   VAR_INPUT
      systemArmed : Bool;
      autoBusy : Bool;
      servBusy : Bool;
      teachingRunning : Bool;
      startUsRunning : Bool;
      modeRequest : UInt;
      modeReqSeq : UInt;
   END_VAR
   VAR_OUTPUT
      modeEffective : UInt;
      modeReady : Bool;
      enterService : Bool;
      enterAuto : Bool;
   END_VAR
   VAR
      lastSeq : UInt;
      safeAllOk : Bool;
      windowAuto : Bool;
      acceptSrv : Bool;
      acceptAuto : Bool;
   END_VAR
BEGIN

REGION Network 1 (SCL)
   #safeAllOk := #systemArmed;
   // Ventana AUTO: OR de todos los *_running (ver tablas por etapa en el PDF).  // nivel sostenido
   #windowAuto :=
   #teachingRunning OR #startUsRunning;

   #enterService := FALSE;
   #enterAuto := FALSE;
   #acceptSrv := FALSE;
   #acceptAuto := FALSE;
END_REGION

REGION Network 2 (SCL)
   // 1) Nueva petición por contador
   IF #modeReqSeq <> #lastSeq THEN
       #lastSeq := #modeReqSeq;

       CASE #modeRequest OF
           0:  // SERVICE
               IF #safeAllOk AND (NOT #autoBusy) AND (NOT #windowAuto) THEN
                   #acceptSrv := TRUE;
               END_IF;

           1:  // AUTO
               IF #safeAllOk AND (NOT #servBusy) THEN
                   #acceptAuto := TRUE;
               END_IF;

       END_CASE;
   END_IF;
END_REGION

REGION Network 3 (SCL)
   IF #acceptSrv THEN
       #modeEffective := 0;
       #enterService := TRUE;
   ELSIF #acceptAuto THEN
       #modeEffective := 1;
       #enterAuto := TRUE;
   END_IF;

   // 3) Ready hacia HMI
   IF #modeEffective = 0 THEN
       #modeReady := #safeAllOk AND (NOT #autoBusy);
   ELSE
       #modeReady := #safeAllOk AND (NOT #servBusy);
   END_IF;
END_REGION
END_FUNCTION_BLOCK

FUNCTION_BLOCK "KukaControlSeq"   // FB21, LAD
{ S7_Optimized_Access := 'TRUE' }
VERSION : 0.1
BEGIN

REGION Network 1: Envia posiciones a la aplicacion KukaControl
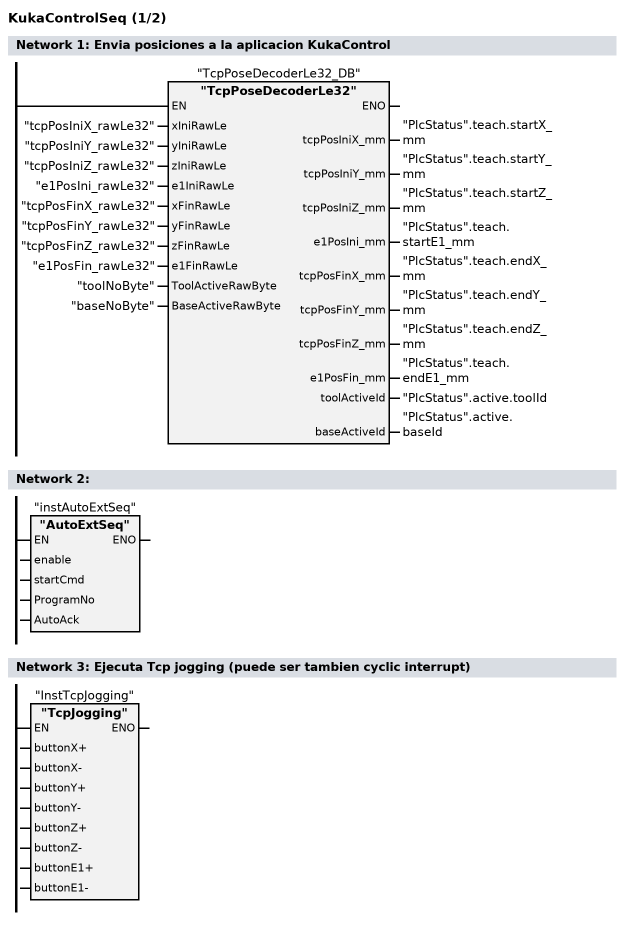
   RUNG wire#powerrail
      "TcpPoseDecoderLe32_DB"(xIniRawLe := "tcpPosIniX_rawLe32", yIniRawLe := "tcpPosIniY_rawLe32", zIniRawLe := "tcpPosIniZ_rawLe32", e1IniRawLe := "e1PosIni_rawLe32", xFinRawLe := "tcpPosFinX_rawLe32", yFinRawLe := "tcpPosFinY_rawLe32", zFinRawLe := "tcpPosFinZ_rawLe32", e1FinRawLe := "e1PosFin_rawLe32", ToolActiveRawByte := "toolNoByte", BaseActiveRawByte := "baseNoByte", tcpPosIniX_mm => "PlcStatus".teach.startX_mm, tcpPosIniY_mm => "PlcStatus".teach.startY_mm, tcpPosIniZ_mm => "PlcStatus".teach.startZ_mm, e1PosIni_mm => "PlcStatus".teach.startE1_mm, tcpPosFinX_mm => "PlcStatus".teach.endX_mm, tcpPosFinY_mm => "PlcStatus".teach.endY_mm, tcpPosFinZ_mm => "PlcStatus".teach.endZ_mm, e1PosFin_mm => "PlcStatus".teach.endE1_mm, toolActiveId => "PlcStatus".active.toolId, baseActiveId => "PlcStatus".active.baseId)
   END_RUNG
   // the same network as SCL:
   "TcpPoseDecoderLe32_DB"(xIniRawLe := "tcpPosIniX_rawLe32",   // "TcpPoseDecoderLe32"
                           yIniRawLe := "tcpPosIniY_rawLe32",
                           zIniRawLe := "tcpPosIniZ_rawLe32",
                           e1IniRawLe := "e1PosIni_rawLe32",
                           xFinRawLe := "tcpPosFinX_rawLe32",
                           yFinRawLe := "tcpPosFinY_rawLe32",
                           zFinRawLe := "tcpPosFinZ_rawLe32",
                           e1FinRawLe := "e1PosFin_rawLe32",
                           ToolActiveRawByte := "toolNoByte",
                           BaseActiveRawByte := "baseNoByte",
                           tcpPosIniX_mm => "PlcStatus".teach.startX_mm,
                           tcpPosIniY_mm => "PlcStatus".teach.startY_mm,
                           tcpPosIniZ_mm => "PlcStatus".teach.startZ_mm,
                           e1PosIni_mm => "PlcStatus".teach.startE1_mm,
                           tcpPosFinX_mm => "PlcStatus".teach.endX_mm,
                           tcpPosFinY_mm => "PlcStatus".teach.endY_mm,
                           tcpPosFinZ_mm => "PlcStatus".teach.endZ_mm,
                           e1PosFin_mm => "PlcStatus".teach.endE1_mm,
                           toolActiveId => "PlcStatus".active.toolId,
                           baseActiveId => "PlcStatus".active.baseId);
END_REGION

REGION Network 2
   RUNG wire#powerrail
      "instAutoExtSeq"(enable :=, startCmd :=, ProgramNo :=, AutoAck :=)
   END_RUNG
   // the same network as SCL:
   "instAutoExtSeq"();   // "AutoExtSeq"
END_REGION

REGION Network 3: Ejecuta Tcp jogging (puede ser tambien cyclic interrupt)
   RUNG wire#powerrail
      "InstTcpJogging"("buttonX+" :=, "buttonX-" :=, "buttonY+" :=, "buttonY-" :=, "buttonZ+" :=, "buttonZ-" :=, "buttonE1+" :=, "buttonE1-" :=)
   END_RUNG
   // the same network as SCL:
   "InstTcpJogging"();   // "TcpJogging"
END_REGION

REGION Network 4: Ejecuta TcpTarget
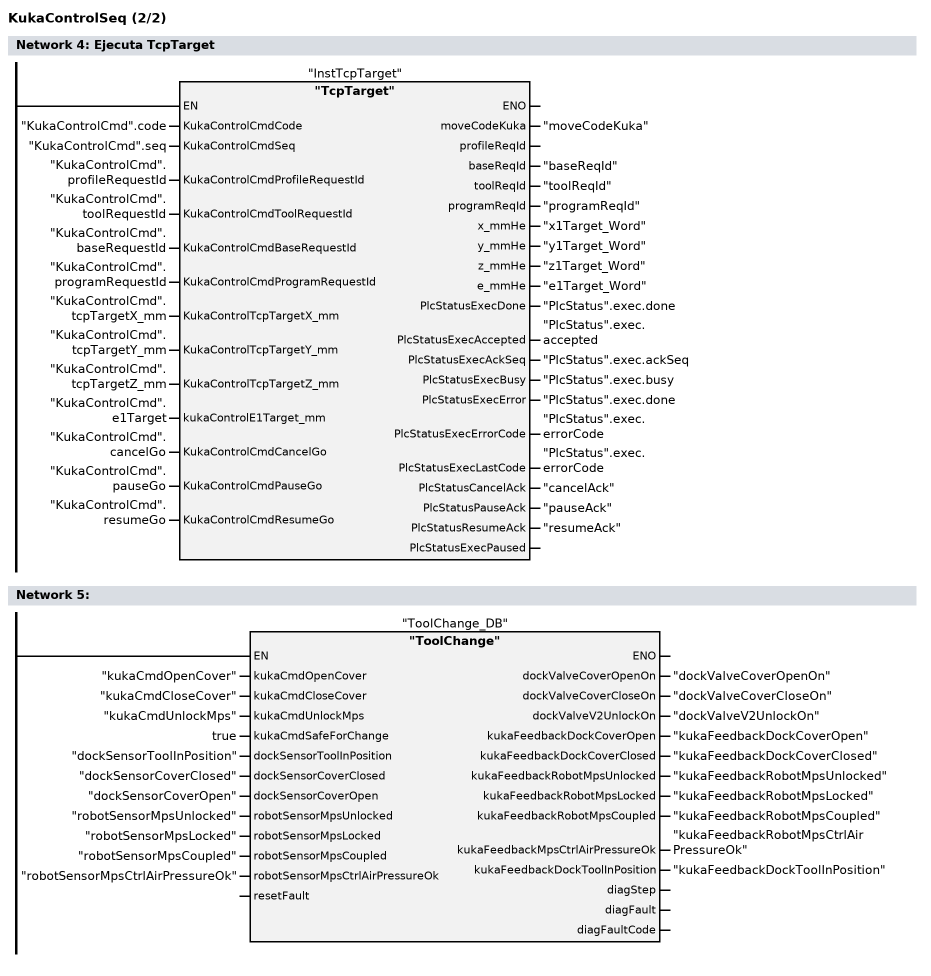
   RUNG wire#powerrail
      "InstTcpTarget"(KukaControlCmdCode := "KukaControlCmd".code, KukaControlCmdSeq := "KukaControlCmd".seq, KukaControlCmdProfileRequestId := "KukaControlCmd".profileRequestId, KukaControlCmdToolRequestId := "KukaControlCmd".toolRequestId, KukaControlCmdBaseRequestId := "KukaControlCmd".baseRequestId, KukaControlCmdProgramRequestId := "KukaControlCmd".programRequestId, KukaControlTcpTargetX_mm := "KukaControlCmd".tcpTargetX_mm, KukaControlTcpTargetY_mm := "KukaControlCmd".tcpTargetY_mm, KukaControlTcpTargetZ_mm := "KukaControlCmd".tcpTargetZ_mm, kukaControlE1Target_mm := "KukaControlCmd".e1Target, KukaControlCmdCancelGo := "KukaControlCmd".cancelGo, KukaControlCmdPauseGo := "KukaControlCmd".pauseGo, KukaControlCmdResumeGo := "KukaControlCmd".resumeGo, moveCodeKuka => "moveCodeKuka", profileReqId =>, baseReqId => "baseReqId", toolReqId => "toolReqId", programReqId => "programReqId", x_mmHe => "x1Target_Word", y_mmHe => "y1Target_Word", z_mmHe => "z1Target_Word", e_mmHe => "e1Target_Word", PlcStatusExecDone => "PlcStatus".exec.done, PlcStatusExecAccepted => "PlcStatus".exec.accepted, PlcStatusExecAckSeq => "PlcStatus".exec.ackSeq, PlcStatusExecBusy => "PlcStatus".exec.busy, PlcStatusExecError => "PlcStatus".exec.done, PlcStatusExecErrorCode => "PlcStatus".exec.errorCode, PlcStatusExecLastCode => "PlcStatus".exec.errorCode, PlcStatusCancelAck => "cancelAck", PlcStatusPauseAck => "pauseAck", PlcStatusResumeAck => "resumeAck", PlcStatusExecPaused =>)
   END_RUNG
   // the same network as SCL:
   "InstTcpTarget"(KukaControlCmdCode := "KukaControlCmd".code,   // "TcpTarget"
                   KukaControlCmdSeq := "KukaControlCmd".seq,
                   KukaControlCmdProfileRequestId := "KukaControlCmd".profileRequestId,
                   KukaControlCmdToolRequestId := "KukaControlCmd".toolRequestId,
                   KukaControlCmdBaseRequestId := "KukaControlCmd".baseRequestId,
                   KukaControlCmdProgramRequestId := "KukaControlCmd".programRequestId,
                   KukaControlTcpTargetX_mm := "KukaControlCmd".tcpTargetX_mm,
                   KukaControlTcpTargetY_mm := "KukaControlCmd".tcpTargetY_mm,
                   KukaControlTcpTargetZ_mm := "KukaControlCmd".tcpTargetZ_mm,
                   kukaControlE1Target_mm := "KukaControlCmd".e1Target,
                   KukaControlCmdCancelGo := "KukaControlCmd".cancelGo,
                   KukaControlCmdPauseGo := "KukaControlCmd".pauseGo,
                   KukaControlCmdResumeGo := "KukaControlCmd".resumeGo,
                   moveCodeKuka => "moveCodeKuka",
                   baseReqId => "baseReqId",
                   toolReqId => "toolReqId",
                   programReqId => "programReqId",
                   x_mmHe => "x1Target_Word",
                   y_mmHe => "y1Target_Word",
                   z_mmHe => "z1Target_Word",
                   e_mmHe => "e1Target_Word",
                   PlcStatusExecDone => "PlcStatus".exec.done,
                   PlcStatusExecAccepted => "PlcStatus".exec.accepted,
                   PlcStatusExecAckSeq => "PlcStatus".exec.ackSeq,
                   PlcStatusExecBusy => "PlcStatus".exec.busy,
                   PlcStatusExecError => "PlcStatus".exec.done,
                   PlcStatusExecErrorCode => "PlcStatus".exec.errorCode,
                   PlcStatusExecLastCode => "PlcStatus".exec.errorCode,
                   PlcStatusCancelAck => "cancelAck",
                   PlcStatusPauseAck => "pauseAck",
                   PlcStatusResumeAck => "resumeAck");
END_REGION
